(* Logix 5000 project; controller MV vendor 1 type 14 code 217 rev 31.11; software revision 31.00; part 48 of 53 *)
(* tags used below, declared in another part *)
   CWD : CHECKWORD_FLAGS;
   Delphi_Does_Eng_Func : BOOL;
   MV_MV1R : PlantItem;   // MV1R
   MV_MV20_CV1 : PlantItem;   // MV20_CV1
   MV_MV21_CV1 : PlantItem;   // MV21_CV1
   MV_MV22_CV1 : PlantItem;   // MV22_CV1
   MV_MV23_CV1 : PlantItem;   // MV23_CV1
   MV_MV2R : PlantItem;   // MV2R
   MV_MV35_CV1 : PlantItem;   // MV35_CV1
   MV_MV36_AV01 : PlantItem;   // MV36_AV01
   MV_MV37_AV01 : PlantItem;   // MV37_AV01
   MV_MV38_AV01 : PlantItem;   // MV38_AV01
   MV_MV39_AV01 : PlantItem;   // MV39_AV01
   MV_MV3R : PlantItem;   // MV3R
   MV_MV40_AV01 : PlantItem;   // MV40_AV01
   MV_MV41_AV01 : PlantItem;   // MV41_AV01
   MV_MV42_AV01 : PlantItem;   // MV42_AV01
   MV_MV43_AV01 : PlantItem;   // MV43_AV01
   MV_MV44_AV01 : PlantItem;   // MV44_AV01
   MV_MV45_AV01 : PlantItem;   // MV45_AV01
   MV_MV46_AV01 : PlantItem;   // MV46_AV01
   MV_MV47_AV01 : PlantItem;   // MV47_AV01
   MV_MV4R : PlantItem;   // MV4R
   MV_MV5R : PlantItem;   // MV5R
   MV_MV6R : PlantItem;   // MV6R
   MV_MV7R : PlantItem;   // MV7R
   MV_N255 : DINT[255];   // Old Format Checkwords To Keep Delphi Indicating Status Correctly.
(* MV_Common, continued *)

   24: [XIC(Delphi_Does_Eng_Func) [[XIC(MV_N255[24].8) [OTL(MV_MV35_CV1.CW.[CWD.MANUAL]) ,XIC(MV_N255[24].9) OTL(MV_MV35_CV1.CW.[CWD.MANDRV]) ,XIO(MV_N255[24].9) OTU(MV_MV35_CV1.CW.[CWD.MANDRV]) ] ,XIO(MV_N255[24].8) [OTU(MV_MV35_CV1.CW.[CWD.MANUAL]) ,[XIC(MV_MV35_CV1.CW.[CWD.OUTPUT]) OTL(MV_N255[24].9) ,XIO(MV_MV35_CV1.CW.[CWD.OUTPUT]) OTU(MV_N255[24].9) ] ] ] ,[XIC(MV_N255[24].13) OTL(MV_MV35_CV1.CW.[CWD.CHECKOFF]) ,XIO(MV_N255[24].13) OTU(MV_MV35_CV1.CW.[CWD.CHECKOFF]) ] ] ,XIO(Delphi_Does_Eng_Func) [[XIC(MV_MV35_CV1.CW.[CWD.MANUAL]) OTL(MV_N255[24].8) ,XIO(MV_MV35_CV1.CW.[CWD.MANUAL]) OTU(MV_N255[24].8) ] ,[XIC(MV_MV35_CV1.CW.[CWD.CHECKOFF]) OTL(MV_N255[24].13) ,XIO(MV_MV35_CV1.CW.[CWD.CHECKOFF]) OTU(MV_N255[24].13) ] ,[XIC(MV_MV35_CV1.CW.[CWD.OUTPUT]) OTL(MV_N255[24].9) ,XIO(MV_MV35_CV1.CW.[CWD.OUTPUT]) OTU(MV_N255[24].9) ] ] ,XIC(MV_MV35_CV1.CW.[CWD.OUTPUT]) OTE(MV_N255[24].10) ,XIO(MV_MV35_CV1.CW.[CWD.OUTPUT]) OTE(MV_N255[24].11) ,XIC(MV_MV35_CV1.CW.[CWD.FAULT]) OTE(MV_N255[24].15) ];
   25: [XIC(Delphi_Does_Eng_Func) [[XIC(MV_N255[25].8) [OTL(MV_MV20_CV1.CW.[CWD.MANUAL]) ,XIC(MV_N255[25].9) OTL(MV_MV20_CV1.CW.[CWD.MANDRV]) ,XIO(MV_N255[25].9) OTU(MV_MV20_CV1.CW.[CWD.MANDRV]) ] ,XIO(MV_N255[25].8) [OTU(MV_MV20_CV1.CW.[CWD.MANUAL]) ,[XIC(MV_MV20_CV1.CW.[CWD.OUTPUT]) OTL(MV_N255[25].9) ,XIO(MV_MV20_CV1.CW.[CWD.OUTPUT]) OTU(MV_N255[25].9) ] ] ] ,[XIC(MV_N255[25].13) OTL(MV_MV20_CV1.CW.[CWD.CHECKOFF]) ,XIO(MV_N255[25].13) OTU(MV_MV20_CV1.CW.[CWD.CHECKOFF]) ] ] ,XIO(Delphi_Does_Eng_Func) [[XIC(MV_MV20_CV1.CW.[CWD.MANUAL]) OTL(MV_N255[25].8) ,XIO(MV_MV20_CV1.CW.[CWD.MANUAL]) OTU(MV_N255[25].8) ] ,[XIC(MV_MV20_CV1.CW.[CWD.CHECKOFF]) OTL(MV_N255[25].13) ,XIO(MV_MV20_CV1.CW.[CWD.CHECKOFF]) OTU(MV_N255[25].13) ] ,[XIC(MV_MV20_CV1.CW.[CWD.OUTPUT]) OTL(MV_N255[25].9) ,XIO(MV_MV20_CV1.CW.[CWD.OUTPUT]) OTU(MV_N255[25].9) ] ] ,XIC(MV_MV20_CV1.CW.[CWD.OUTPUT]) OTE(MV_N255[25].10) ,XIO(MV_MV20_CV1.CW.[CWD.OUTPUT]) OTE(MV_N255[25].11) ,XIC(MV_MV20_CV1.CW.[CWD.FAULT]) OTE(MV_N255[25].15) ];
   26: [XIC(Delphi_Does_Eng_Func) [[XIC(MV_N255[26].8) [OTL(MV_MV21_CV1.CW.[CWD.MANUAL]) ,XIC(MV_N255[26].9) OTL(MV_MV21_CV1.CW.[CWD.MANDRV]) ,XIO(MV_N255[26].9) OTU(MV_MV21_CV1.CW.[CWD.MANDRV]) ] ,XIO(MV_N255[26].8) [OTU(MV_MV21_CV1.CW.[CWD.MANUAL]) ,[XIC(MV_MV21_CV1.CW.[CWD.OUTPUT]) OTL(MV_N255[26].9) ,XIO(MV_MV21_CV1.CW.[CWD.OUTPUT]) OTU(MV_N255[26].9) ] ] ] ,[XIC(MV_N255[26].13) OTL(MV_MV21_CV1.CW.[CWD.CHECKOFF]) ,XIO(MV_N255[26].13) OTU(MV_MV21_CV1.CW.[CWD.CHECKOFF]) ] ] ,XIO(Delphi_Does_Eng_Func) [[XIC(MV_MV21_CV1.CW.[CWD.MANUAL]) OTL(MV_N255[26].8) ,XIO(MV_MV21_CV1.CW.[CWD.MANUAL]) OTU(MV_N255[26].8) ] ,[XIC(MV_MV21_CV1.CW.[CWD.CHECKOFF]) OTL(MV_N255[26].13) ,XIO(MV_MV21_CV1.CW.[CWD.CHECKOFF]) OTU(MV_N255[26].13) ] ,[XIC(MV_MV21_CV1.CW.[CWD.OUTPUT]) OTL(MV_N255[26].9) ,XIO(MV_MV21_CV1.CW.[CWD.OUTPUT]) OTU(MV_N255[26].9) ] ] ,XIC(MV_MV21_CV1.CW.[CWD.OUTPUT]) OTE(MV_N255[26].10) ,XIO(MV_MV21_CV1.CW.[CWD.OUTPUT]) OTE(MV_N255[26].11) ,XIC(MV_MV21_CV1.CW.[CWD.FAULT]) OTE(MV_N255[26].15) ];
   27: [XIC(Delphi_Does_Eng_Func) [[XIC(MV_N255[27].8) [OTL(MV_MV22_CV1.CW.[CWD.MANUAL]) ,XIC(MV_N255[27].9) OTL(MV_MV22_CV1.CW.[CWD.MANDRV]) ,XIO(MV_N255[27].9) OTU(MV_MV22_CV1.CW.[CWD.MANDRV]) ] ,XIO(MV_N255[27].8) [OTU(MV_MV22_CV1.CW.[CWD.MANUAL]) ,[XIC(MV_MV22_CV1.CW.[CWD.OUTPUT]) OTL(MV_N255[27].9) ,XIO(MV_MV22_CV1.CW.[CWD.OUTPUT]) OTU(MV_N255[27].9) ] ] ] ,[XIC(MV_N255[27].13) OTL(MV_MV22_CV1.CW.[CWD.CHECKOFF]) ,XIO(MV_N255[27].13) OTU(MV_MV22_CV1.CW.[CWD.CHECKOFF]) ] ] ,XIO(Delphi_Does_Eng_Func) [[XIC(MV_MV22_CV1.CW.[CWD.MANUAL]) OTL(MV_N255[27].8) ,XIO(MV_MV22_CV1.CW.[CWD.MANUAL]) OTU(MV_N255[27].8) ] ,[XIC(MV_MV22_CV1.CW.[CWD.CHECKOFF]) OTL(MV_N255[27].13) ,XIO(MV_MV22_CV1.CW.[CWD.CHECKOFF]) OTU(MV_N255[27].13) ] ,[XIC(MV_MV22_CV1.CW.[CWD.OUTPUT]) OTL(MV_N255[27].9) ,XIO(MV_MV22_CV1.CW.[CWD.OUTPUT]) OTU(MV_N255[27].9) ] ] ,XIC(MV_MV22_CV1.CW.[CWD.OUTPUT]) OTE(MV_N255[27].10) ,XIO(MV_MV22_CV1.CW.[CWD.OUTPUT]) OTE(MV_N255[27].11) ,XIC(MV_MV22_CV1.CW.[CWD.FAULT]) OTE(MV_N255[27].15) ];
   28: [XIC(Delphi_Does_Eng_Func) [[XIC(MV_N255[28].8) [OTL(MV_MV23_CV1.CW.[CWD.MANUAL]) ,XIC(MV_N255[28].9) OTL(MV_MV23_CV1.CW.[CWD.MANDRV]) ,XIO(MV_N255[28].9) OTU(MV_MV23_CV1.CW.[CWD.MANDRV]) ] ,XIO(MV_N255[28].8) [OTU(MV_MV23_CV1.CW.[CWD.MANUAL]) ,[XIC(MV_MV23_CV1.CW.[CWD.OUTPUT]) OTL(MV_N255[28].9) ,XIO(MV_MV23_CV1.CW.[CWD.OUTPUT]) OTU(MV_N255[28].9) ] ] ] ,[XIC(MV_N255[28].13) OTL(MV_MV23_CV1.CW.[CWD.CHECKOFF]) ,XIO(MV_N255[28].13) OTU(MV_MV23_CV1.CW.[CWD.CHECKOFF]) ] ] ,XIO(Delphi_Does_Eng_Func) [[XIC(MV_MV23_CV1.CW.[CWD.MANUAL]) OTL(MV_N255[28].8) ,XIO(MV_MV23_CV1.CW.[CWD.MANUAL]) OTU(MV_N255[28].8) ] ,[XIC(MV_MV23_CV1.CW.[CWD.CHECKOFF]) OTL(MV_N255[28].13) ,XIO(MV_MV23_CV1.CW.[CWD.CHECKOFF]) OTU(MV_N255[28].13) ] ,[XIC(MV_MV23_CV1.CW.[CWD.OUTPUT]) OTL(MV_N255[28].9) ,XIO(MV_MV23_CV1.CW.[CWD.OUTPUT]) OTU(MV_N255[28].9) ] ] ,XIC(MV_MV23_CV1.CW.[CWD.OUTPUT]) OTE(MV_N255[28].10) ,XIO(MV_MV23_CV1.CW.[CWD.OUTPUT]) OTE(MV_N255[28].11) ,XIC(MV_MV23_CV1.CW.[CWD.FAULT]) OTE(MV_N255[28].15) ];
   29: [XIC(Delphi_Does_Eng_Func) [[XIC(MV_N255[64].8) [OTL(MV_MV36_AV01.CW.[CWD.MANUAL]) ,XIC(MV_N255[64].9) OTL(MV_MV36_AV01.CW.[CWD.MANDRV]) ,XIO(MV_N255[64].9) OTU(MV_MV36_AV01.CW.[CWD.MANDRV]) ] ,XIO(MV_N255[64].8) [OTU(MV_MV36_AV01.CW.[CWD.MANUAL]) ,[XIC(MV_MV36_AV01.CW.[CWD.OUTPUT]) OTL(MV_N255[64].9) ,XIO(MV_MV36_AV01.CW.[CWD.OUTPUT]) OTU(MV_N255[64].9) ] ] ] ,[XIC(MV_N255[64].13) OTL(MV_MV36_AV01.CW.[CWD.CHECKOFF]) ,XIO(MV_N255[64].13) OTU(MV_MV36_AV01.CW.[CWD.CHECKOFF]) ] ] ,XIO(Delphi_Does_Eng_Func) [[XIC(MV_MV36_AV01.CW.[CWD.MANUAL]) OTL(MV_N255[64].8) ,XIO(MV_MV36_AV01.CW.[CWD.MANUAL]) OTU(MV_N255[64].8) ] ,[XIC(MV_MV36_AV01.CW.[CWD.CHECKOFF]) OTL(MV_N255[64].13) ,XIO(MV_MV36_AV01.CW.[CWD.CHECKOFF]) OTU(MV_N255[64].13) ] ,[XIC(MV_MV36_AV01.CW.[CWD.OUTPUT]) OTL(MV_N255[64].9) ,XIO(MV_MV36_AV01.CW.[CWD.OUTPUT]) OTU(MV_N255[64].9) ] ] ,XIC(MV_MV36_AV01.CW.[CWD.OUTPUT]) OTE(MV_N255[64].10) ,XIO(MV_MV36_AV01.CW.[CWD.OUTPUT]) OTE(MV_N255[64].11) ,XIC(MV_MV36_AV01.CW.[CWD.FAULT]) OTE(MV_N255[64].15) ];
   30: [XIC(Delphi_Does_Eng_Func) [[XIC(MV_N255[65].8) [OTL(MV_MV37_AV01.CW.[CWD.MANUAL]) ,XIC(MV_N255[65].9) OTL(MV_MV37_AV01.CW.[CWD.MANDRV]) ,XIO(MV_N255[65].9) OTU(MV_MV37_AV01.CW.[CWD.MANDRV]) ] ,XIO(MV_N255[65].8) [OTU(MV_MV37_AV01.CW.[CWD.MANUAL]) ,[XIC(MV_MV37_AV01.CW.[CWD.OUTPUT]) OTL(MV_N255[65].9) ,XIO(MV_MV37_AV01.CW.[CWD.OUTPUT]) OTU(MV_N255[65].9) ] ] ] ,[XIC(MV_N255[65].13) OTL(MV_MV37_AV01.CW.[CWD.CHECKOFF]) ,XIO(MV_N255[65].13) OTU(MV_MV37_AV01.CW.[CWD.CHECKOFF]) ] ] ,XIO(Delphi_Does_Eng_Func) [[XIC(MV_MV37_AV01.CW.[CWD.MANUAL]) OTL(MV_N255[65].8) ,XIO(MV_MV37_AV01.CW.[CWD.MANUAL]) OTU(MV_N255[65].8) ] ,[XIC(MV_MV37_AV01.CW.[CWD.CHECKOFF]) OTL(MV_N255[65].13) ,XIO(MV_MV37_AV01.CW.[CWD.CHECKOFF]) OTU(MV_N255[65].13) ] ,[XIC(MV_MV37_AV01.CW.[CWD.OUTPUT]) OTL(MV_N255[65].9) ,XIO(MV_MV37_AV01.CW.[CWD.OUTPUT]) OTU(MV_N255[65].9) ] ] ,XIC(MV_MV37_AV01.CW.[CWD.OUTPUT]) OTE(MV_N255[65].10) ,XIO(MV_MV37_AV01.CW.[CWD.OUTPUT]) OTE(MV_N255[65].11) ,XIC(MV_MV37_AV01.CW.[CWD.FAULT]) OTE(MV_N255[65].15) ];
   31: [XIC(Delphi_Does_Eng_Func) [[XIC(MV_N255[66].8) [OTL(MV_MV38_AV01.CW.[CWD.MANUAL]) ,XIC(MV_N255[66].9) OTL(MV_MV38_AV01.CW.[CWD.MANDRV]) ,XIO(MV_N255[66].9) OTU(MV_MV38_AV01.CW.[CWD.MANDRV]) ] ,XIO(MV_N255[66].8) [OTU(MV_MV38_AV01.CW.[CWD.MANUAL]) ,[XIC(MV_MV38_AV01.CW.[CWD.OUTPUT]) OTL(MV_N255[66].9) ,XIO(MV_MV38_AV01.CW.[CWD.OUTPUT]) OTU(MV_N255[66].9) ] ] ] ,[XIC(MV_N255[66].13) OTL(MV_MV38_AV01.CW.[CWD.CHECKOFF]) ,XIO(MV_N255[66].13) OTU(MV_MV38_AV01.CW.[CWD.CHECKOFF]) ] ] ,XIO(Delphi_Does_Eng_Func) [[XIC(MV_MV38_AV01.CW.[CWD.MANUAL]) OTL(MV_N255[66].8) ,XIO(MV_MV38_AV01.CW.[CWD.MANUAL]) OTU(MV_N255[66].8) ] ,[XIC(MV_MV38_AV01.CW.[CWD.CHECKOFF]) OTL(MV_N255[66].13) ,XIO(MV_MV38_AV01.CW.[CWD.CHECKOFF]) OTU(MV_N255[66].13) ] ,[XIC(MV_MV38_AV01.CW.[CWD.OUTPUT]) OTL(MV_N255[66].9) ,XIO(MV_MV38_AV01.CW.[CWD.OUTPUT]) OTU(MV_N255[66].9) ] ] ,XIC(MV_MV38_AV01.CW.[CWD.OUTPUT]) OTE(MV_N255[66].10) ,XIO(MV_MV38_AV01.CW.[CWD.OUTPUT]) OTE(MV_N255[66].11) ,XIC(MV_MV38_AV01.CW.[CWD.FAULT]) OTE(MV_N255[66].15) ];
   32: [XIC(Delphi_Does_Eng_Func) [[XIC(MV_N255[67].8) [OTL(MV_MV39_AV01.CW.[CWD.MANUAL]) ,XIC(MV_N255[67].9) OTL(MV_MV39_AV01.CW.[CWD.MANDRV]) ,XIO(MV_N255[67].9) OTU(MV_MV39_AV01.CW.[CWD.MANDRV]) ] ,XIO(MV_N255[67].8) [OTU(MV_MV39_AV01.CW.[CWD.MANUAL]) ,[XIC(MV_MV39_AV01.CW.[CWD.OUTPUT]) OTL(MV_N255[67].9) ,XIO(MV_MV39_AV01.CW.[CWD.OUTPUT]) OTU(MV_N255[67].9) ] ] ] ,[XIC(MV_N255[67].13) OTL(MV_MV39_AV01.CW.[CWD.CHECKOFF]) ,XIO(MV_N255[67].13) OTU(MV_MV39_AV01.CW.[CWD.CHECKOFF]) ] ] ,XIO(Delphi_Does_Eng_Func) [[XIC(MV_MV39_AV01.CW.[CWD.MANUAL]) OTL(MV_N255[67].8) ,XIO(MV_MV39_AV01.CW.[CWD.MANUAL]) OTU(MV_N255[67].8) ] ,[XIC(MV_MV39_AV01.CW.[CWD.CHECKOFF]) OTL(MV_N255[67].13) ,XIO(MV_MV39_AV01.CW.[CWD.CHECKOFF]) OTU(MV_N255[67].13) ] ,[XIC(MV_MV39_AV01.CW.[CWD.OUTPUT]) OTL(MV_N255[67].9) ,XIO(MV_MV39_AV01.CW.[CWD.OUTPUT]) OTU(MV_N255[67].9) ] ] ,XIC(MV_MV39_AV01.CW.[CWD.OUTPUT]) OTE(MV_N255[67].10) ,XIO(MV_MV39_AV01.CW.[CWD.OUTPUT]) OTE(MV_N255[67].11) ,XIC(MV_MV39_AV01.CW.[CWD.FAULT]) OTE(MV_N255[67].15) ];
   33: [XIC(Delphi_Does_Eng_Func) [[XIC(MV_N255[68].8) [OTL(MV_MV40_AV01.CW.[CWD.MANUAL]) ,XIC(MV_N255[68].9) OTL(MV_MV40_AV01.CW.[CWD.MANDRV]) ,XIO(MV_N255[68].9) OTU(MV_MV40_AV01.CW.[CWD.MANDRV]) ] ,XIO(MV_N255[68].8) [OTU(MV_MV40_AV01.CW.[CWD.MANUAL]) ,[XIC(MV_MV40_AV01.CW.[CWD.OUTPUT]) OTL(MV_N255[68].9) ,XIO(MV_MV40_AV01.CW.[CWD.OUTPUT]) OTU(MV_N255[68].9) ] ] ] ,[XIC(MV_N255[68].13) OTL(MV_MV40_AV01.CW.[CWD.CHECKOFF]) ,XIO(MV_N255[68].13) OTU(MV_MV40_AV01.CW.[CWD.CHECKOFF]) ] ] ,XIO(Delphi_Does_Eng_Func) [[XIC(MV_MV40_AV01.CW.[CWD.MANUAL]) OTL(MV_N255[68].8) ,XIO(MV_MV40_AV01.CW.[CWD.MANUAL]) OTU(MV_N255[68].8) ] ,[XIC(MV_MV40_AV01.CW.[CWD.CHECKOFF]) OTL(MV_N255[68].13) ,XIO(MV_MV40_AV01.CW.[CWD.CHECKOFF]) OTU(MV_N255[68].13) ] ,[XIC(MV_MV40_AV01.CW.[CWD.OUTPUT]) OTL(MV_N255[68].9) ,XIO(MV_MV40_AV01.CW.[CWD.OUTPUT]) OTU(MV_N255[68].9) ] ] ,XIC(MV_MV40_AV01.CW.[CWD.OUTPUT]) OTE(MV_N255[68].10) ,XIO(MV_MV40_AV01.CW.[CWD.OUTPUT]) OTE(MV_N255[68].11) ,XIC(MV_MV40_AV01.CW.[CWD.FAULT]) OTE(MV_N255[68].15) ];
   34: [XIC(Delphi_Does_Eng_Func) [[XIC(MV_N255[69].8) [OTL(MV_MV41_AV01.CW.[CWD.MANUAL]) ,XIC(MV_N255[69].9) OTL(MV_MV41_AV01.CW.[CWD.MANDRV]) ,XIO(MV_N255[69].9) OTU(MV_MV41_AV01.CW.[CWD.MANDRV]) ] ,XIO(MV_N255[69].8) [OTU(MV_MV41_AV01.CW.[CWD.MANUAL]) ,[XIC(MV_MV41_AV01.CW.[CWD.OUTPUT]) OTL(MV_N255[69].9) ,XIO(MV_MV41_AV01.CW.[CWD.OUTPUT]) OTU(MV_N255[69].9) ] ] ] ,[XIC(MV_N255[69].13) OTL(MV_MV41_AV01.CW.[CWD.CHECKOFF]) ,XIO(MV_N255[69].13) OTU(MV_MV41_AV01.CW.[CWD.CHECKOFF]) ] ] ,XIO(Delphi_Does_Eng_Func) [[XIC(MV_MV41_AV01.CW.[CWD.MANUAL]) OTL(MV_N255[69].8) ,XIO(MV_MV41_AV01.CW.[CWD.MANUAL]) OTU(MV_N255[69].8) ] ,[XIC(MV_MV41_AV01.CW.[CWD.CHECKOFF]) OTL(MV_N255[69].13) ,XIO(MV_MV41_AV01.CW.[CWD.CHECKOFF]) OTU(MV_N255[69].13) ] ,[XIC(MV_MV41_AV01.CW.[CWD.OUTPUT]) OTL(MV_N255[69].9) ,XIO(MV_MV41_AV01.CW.[CWD.OUTPUT]) OTU(MV_N255[69].9) ] ] ,XIC(MV_MV41_AV01.CW.[CWD.OUTPUT]) OTE(MV_N255[69].10) ,XIO(MV_MV41_AV01.CW.[CWD.OUTPUT]) OTE(MV_N255[69].11) ,XIC(MV_MV41_AV01.CW.[CWD.FAULT]) OTE(MV_N255[69].15) ];
   35: [XIC(Delphi_Does_Eng_Func) [[XIC(MV_N255[70].8) [OTL(MV_MV42_AV01.CW.[CWD.MANUAL]) ,XIC(MV_N255[70].9) OTL(MV_MV42_AV01.CW.[CWD.MANDRV]) ,XIO(MV_N255[70].9) OTU(MV_MV42_AV01.CW.[CWD.MANDRV]) ] ,XIO(MV_N255[70].8) [OTU(MV_MV42_AV01.CW.[CWD.MANUAL]) ,[XIC(MV_MV42_AV01.CW.[CWD.OUTPUT]) OTL(MV_N255[70].9) ,XIO(MV_MV42_AV01.CW.[CWD.OUTPUT]) OTU(MV_N255[70].9) ] ] ] ,[XIC(MV_N255[70].13) OTL(MV_MV42_AV01.CW.[CWD.CHECKOFF]) ,XIO(MV_N255[70].13) OTU(MV_MV42_AV01.CW.[CWD.CHECKOFF]) ] ] ,XIO(Delphi_Does_Eng_Func) [[XIC(MV_MV42_AV01.CW.[CWD.MANUAL]) OTL(MV_N255[70].8) ,XIO(MV_MV42_AV01.CW.[CWD.MANUAL]) OTU(MV_N255[70].8) ] ,[XIC(MV_MV42_AV01.CW.[CWD.CHECKOFF]) OTL(MV_N255[70].13) ,XIO(MV_MV42_AV01.CW.[CWD.CHECKOFF]) OTU(MV_N255[70].13) ] ,[XIC(MV_MV42_AV01.CW.[CWD.OUTPUT]) OTL(MV_N255[70].9) ,XIO(MV_MV42_AV01.CW.[CWD.OUTPUT]) OTU(MV_N255[70].9) ] ] ,XIC(MV_MV42_AV01.CW.[CWD.OUTPUT]) OTE(MV_N255[70].10) ,XIO(MV_MV42_AV01.CW.[CWD.OUTPUT]) OTE(MV_N255[70].11) ,XIC(MV_MV42_AV01.CW.[CWD.FAULT]) OTE(MV_N255[70].15) ];
   36: [XIC(Delphi_Does_Eng_Func) [[XIC(MV_N255[71].8) [OTL(MV_MV43_AV01.CW.[CWD.MANUAL]) ,XIC(MV_N255[71].9) OTL(MV_MV43_AV01.CW.[CWD.MANDRV]) ,XIO(MV_N255[71].9) OTU(MV_MV43_AV01.CW.[CWD.MANDRV]) ] ,XIO(MV_N255[71].8) [OTU(MV_MV43_AV01.CW.[CWD.MANUAL]) ,[XIC(MV_MV43_AV01.CW.[CWD.OUTPUT]) OTL(MV_N255[71].9) ,XIO(MV_MV43_AV01.CW.[CWD.OUTPUT]) OTU(MV_N255[71].9) ] ] ] ,[XIC(MV_N255[71].13) OTL(MV_MV43_AV01.CW.[CWD.CHECKOFF]) ,XIO(MV_N255[71].13) OTU(MV_MV43_AV01.CW.[CWD.CHECKOFF]) ] ] ,XIO(Delphi_Does_Eng_Func) [[XIC(MV_MV43_AV01.CW.[CWD.MANUAL]) OTL(MV_N255[71].8) ,XIO(MV_MV43_AV01.CW.[CWD.MANUAL]) OTU(MV_N255[71].8) ] ,[XIC(MV_MV43_AV01.CW.[CWD.CHECKOFF]) OTL(MV_N255[71].13) ,XIO(MV_MV43_AV01.CW.[CWD.CHECKOFF]) OTU(MV_N255[71].13) ] ,[XIC(MV_MV43_AV01.CW.[CWD.OUTPUT]) OTL(MV_N255[71].9) ,XIO(MV_MV43_AV01.CW.[CWD.OUTPUT]) OTU(MV_N255[71].9) ] ] ,XIC(MV_MV43_AV01.CW.[CWD.OUTPUT]) OTE(MV_N255[71].10) ,XIO(MV_MV43_AV01.CW.[CWD.OUTPUT]) OTE(MV_N255[71].11) ,XIC(MV_MV43_AV01.CW.[CWD.FAULT]) OTE(MV_N255[71].15) ];
   37: [XIC(Delphi_Does_Eng_Func) [[XIC(MV_N255[72].8) [OTL(MV_MV44_AV01.CW.[CWD.MANUAL]) ,XIC(MV_N255[72].9) OTL(MV_MV44_AV01.CW.[CWD.MANDRV]) ,XIO(MV_N255[72].9) OTU(MV_MV44_AV01.CW.[CWD.MANDRV]) ] ,XIO(MV_N255[72].8) [OTU(MV_MV44_AV01.CW.[CWD.MANUAL]) ,[XIC(MV_MV44_AV01.CW.[CWD.OUTPUT]) OTL(MV_N255[72].9) ,XIO(MV_MV44_AV01.CW.[CWD.OUTPUT]) OTU(MV_N255[72].9) ] ] ] ,[XIC(MV_N255[72].13) OTL(MV_MV44_AV01.CW.[CWD.CHECKOFF]) ,XIO(MV_N255[72].13) OTU(MV_MV44_AV01.CW.[CWD.CHECKOFF]) ] ] ,XIO(Delphi_Does_Eng_Func) [[XIC(MV_MV44_AV01.CW.[CWD.MANUAL]) OTL(MV_N255[72].8) ,XIO(MV_MV44_AV01.CW.[CWD.MANUAL]) OTU(MV_N255[72].8) ] ,[XIC(MV_MV44_AV01.CW.[CWD.CHECKOFF]) OTL(MV_N255[72].13) ,XIO(MV_MV44_AV01.CW.[CWD.CHECKOFF]) OTU(MV_N255[72].13) ] ,[XIC(MV_MV44_AV01.CW.[CWD.OUTPUT]) OTL(MV_N255[72].9) ,XIO(MV_MV44_AV01.CW.[CWD.OUTPUT]) OTU(MV_N255[72].9) ] ] ,XIC(MV_MV44_AV01.CW.[CWD.OUTPUT]) OTE(MV_N255[72].10) ,XIO(MV_MV44_AV01.CW.[CWD.OUTPUT]) OTE(MV_N255[72].11) ,XIC(MV_MV44_AV01.CW.[CWD.FAULT]) OTE(MV_N255[72].15) ];
   38: [XIC(Delphi_Does_Eng_Func) [[XIC(MV_N255[73].8) [OTL(MV_MV45_AV01.CW.[CWD.MANUAL]) ,XIC(MV_N255[73].9) OTL(MV_MV45_AV01.CW.[CWD.MANDRV]) ,XIO(MV_N255[73].9) OTU(MV_MV45_AV01.CW.[CWD.MANDRV]) ] ,XIO(MV_N255[73].8) [OTU(MV_MV45_AV01.CW.[CWD.MANUAL]) ,[XIC(MV_MV45_AV01.CW.[CWD.OUTPUT]) OTL(MV_N255[73].9) ,XIO(MV_MV45_AV01.CW.[CWD.OUTPUT]) OTU(MV_N255[73].9) ] ] ] ,[XIC(MV_N255[73].13) OTL(MV_MV45_AV01.CW.[CWD.CHECKOFF]) ,XIO(MV_N255[73].13) OTU(MV_MV45_AV01.CW.[CWD.CHECKOFF]) ] ] ,XIO(Delphi_Does_Eng_Func) [[XIC(MV_MV45_AV01.CW.[CWD.MANUAL]) OTL(MV_N255[73].8) ,XIO(MV_MV45_AV01.CW.[CWD.MANUAL]) OTU(MV_N255[73].8) ] ,[XIC(MV_MV45_AV01.CW.[CWD.CHECKOFF]) OTL(MV_N255[73].13) ,XIO(MV_MV45_AV01.CW.[CWD.CHECKOFF]) OTU(MV_N255[73].13) ] ,[XIC(MV_MV45_AV01.CW.[CWD.OUTPUT]) OTL(MV_N255[73].9) ,XIO(MV_MV45_AV01.CW.[CWD.OUTPUT]) OTU(MV_N255[73].9) ] ] ,XIC(MV_MV45_AV01.CW.[CWD.OUTPUT]) OTE(MV_N255[73].10) ,XIO(MV_MV45_AV01.CW.[CWD.OUTPUT]) OTE(MV_N255[73].11) ,XIC(MV_MV45_AV01.CW.[CWD.FAULT]) OTE(MV_N255[73].15) ];
   39: [XIC(Delphi_Does_Eng_Func) [[XIC(MV_N255[74].8) [OTL(MV_MV46_AV01.CW.[CWD.MANUAL]) ,XIC(MV_N255[74].9) OTL(MV_MV46_AV01.CW.[CWD.MANDRV]) ,XIO(MV_N255[74].9) OTU(MV_MV46_AV01.CW.[CWD.MANDRV]) ] ,XIO(MV_N255[74].8) [OTU(MV_MV46_AV01.CW.[CWD.MANUAL]) ,[XIC(MV_MV46_AV01.CW.[CWD.OUTPUT]) OTL(MV_N255[74].9) ,XIO(MV_MV46_AV01.CW.[CWD.OUTPUT]) OTU(MV_N255[74].9) ] ] ] ,[XIC(MV_N255[74].13) OTL(MV_MV46_AV01.CW.[CWD.CHECKOFF]) ,XIO(MV_N255[74].13) OTU(MV_MV46_AV01.CW.[CWD.CHECKOFF]) ] ] ,XIO(Delphi_Does_Eng_Func) [[XIC(MV_MV46_AV01.CW.[CWD.MANUAL]) OTL(MV_N255[74].8) ,XIO(MV_MV46_AV01.CW.[CWD.MANUAL]) OTU(MV_N255[74].8) ] ,[XIC(MV_MV46_AV01.CW.[CWD.CHECKOFF]) OTL(MV_N255[74].13) ,XIO(MV_MV46_AV01.CW.[CWD.CHECKOFF]) OTU(MV_N255[74].13) ] ,[XIC(MV_MV46_AV01.CW.[CWD.OUTPUT]) OTL(MV_N255[74].9) ,XIO(MV_MV46_AV01.CW.[CWD.OUTPUT]) OTU(MV_N255[74].9) ] ] ,XIC(MV_MV46_AV01.CW.[CWD.OUTPUT]) OTE(MV_N255[74].10) ,XIO(MV_MV46_AV01.CW.[CWD.OUTPUT]) OTE(MV_N255[74].11) ,XIC(MV_MV46_AV01.CW.[CWD.FAULT]) OTE(MV_N255[74].15) ];
   40: [XIC(Delphi_Does_Eng_Func) [[XIC(MV_N255[75].8) [OTL(MV_MV47_AV01.CW.[CWD.MANUAL]) ,XIC(MV_N255[75].9) OTL(MV_MV47_AV01.CW.[CWD.MANDRV]) ,XIO(MV_N255[75].9) OTU(MV_MV47_AV01.CW.[CWD.MANDRV]) ] ,XIO(MV_N255[75].8) [OTU(MV_MV47_AV01.CW.[CWD.MANUAL]) ,[XIC(MV_MV47_AV01.CW.[CWD.OUTPUT]) OTL(MV_N255[75].9) ,XIO(MV_MV47_AV01.CW.[CWD.OUTPUT]) OTU(MV_N255[75].9) ] ] ] ,[XIC(MV_N255[75].13) OTL(MV_MV47_AV01.CW.[CWD.CHECKOFF]) ,XIO(MV_N255[75].13) OTU(MV_MV47_AV01.CW.[CWD.CHECKOFF]) ] ] ,XIO(Delphi_Does_Eng_Func) [[XIC(MV_MV47_AV01.CW.[CWD.MANUAL]) OTL(MV_N255[75].8) ,XIO(MV_MV47_AV01.CW.[CWD.MANUAL]) OTU(MV_N255[75].8) ] ,[XIC(MV_MV47_AV01.CW.[CWD.CHECKOFF]) OTL(MV_N255[75].13) ,XIO(MV_MV47_AV01.CW.[CWD.CHECKOFF]) OTU(MV_N255[75].13) ] ,[XIC(MV_MV47_AV01.CW.[CWD.OUTPUT]) OTL(MV_N255[75].9) ,XIO(MV_MV47_AV01.CW.[CWD.OUTPUT]) OTU(MV_N255[75].9) ] ] ,XIC(MV_MV47_AV01.CW.[CWD.OUTPUT]) OTE(MV_N255[75].10) ,XIO(MV_MV47_AV01.CW.[CWD.OUTPUT]) OTE(MV_N255[75].11) ,XIC(MV_MV47_AV01.CW.[CWD.FAULT]) OTE(MV_N255[75].15) ];
   41: [XIC(Delphi_Does_Eng_Func) [[XIC(MV_N255[32].8) [OTL(MV_MV1R.CW.[CWD.MANUAL]) ,XIC(MV_N255[32].9) OTL(MV_MV1R.CW.[CWD.MANDRV]) ,XIO(MV_N255[32].9) OTU(MV_MV1R.CW.[CWD.MANDRV]) ] ,XIO(MV_N255[32].8) [OTU(MV_MV1R.CW.[CWD.MANUAL]) ,[XIC(MV_MV1R.CW.[CWD.OUTPUT]) OTL(MV_N255[32].9) ,XIO(MV_MV1R.CW.[CWD.OUTPUT]) OTU(MV_N255[32].9) ] ] ] ,[XIC(MV_N255[32].13) OTL(MV_MV1R.CW.[CWD.CHECKOFF]) ,XIO(MV_N255[32].13) OTU(MV_MV1R.CW.[CWD.CHECKOFF]) ] ] ,XIO(Delphi_Does_Eng_Func) [[XIC(MV_MV1R.CW.[CWD.MANUAL]) OTL(MV_N255[32].8) ,XIO(MV_MV1R.CW.[CWD.MANUAL]) OTU(MV_N255[32].8) ] ,[XIC(MV_MV1R.CW.[CWD.CHECKOFF]) OTL(MV_N255[32].13) ,XIO(MV_MV1R.CW.[CWD.CHECKOFF]) OTU(MV_N255[32].13) ] ,[XIC(MV_MV1R.CW.[CWD.OUTPUT]) OTL(MV_N255[32].9) ,XIO(MV_MV1R.CW.[CWD.OUTPUT]) OTU(MV_N255[32].9) ] ] ,XIC(MV_MV1R.CW.[CWD.RUNFB]) OTE(MV_N255[32].10) ,XIO(MV_MV1R.CW.[CWD.RUNFB]) OTE(MV_N255[32].11) ,XIC(MV_MV1R.CW.[CWD.FAULT]) OTE(MV_N255[32].15) ];
   42: [XIC(Delphi_Does_Eng_Func) [[XIC(MV_N255[33].8) [OTL(MV_MV2R.CW.[CWD.MANUAL]) ,XIC(MV_N255[33].9) OTL(MV_MV2R.CW.[CWD.MANDRV]) ,XIO(MV_N255[33].9) OTU(MV_MV2R.CW.[CWD.MANDRV]) ] ,XIO(MV_N255[33].8) [OTU(MV_MV2R.CW.[CWD.MANUAL]) ,[XIC(MV_MV2R.CW.[CWD.OUTPUT]) OTL(MV_N255[33].9) ,XIO(MV_MV2R.CW.[CWD.OUTPUT]) OTU(MV_N255[33].9) ] ] ] ,[XIC(MV_N255[33].13) OTL(MV_MV2R.CW.[CWD.CHECKOFF]) ,XIO(MV_N255[33].13) OTU(MV_MV2R.CW.[CWD.CHECKOFF]) ] ] ,XIO(Delphi_Does_Eng_Func) [[XIC(MV_MV2R.CW.[CWD.MANUAL]) OTL(MV_N255[33].8) ,XIO(MV_MV2R.CW.[CWD.MANUAL]) OTU(MV_N255[33].8) ] ,[XIC(MV_MV2R.CW.[CWD.CHECKOFF]) OTL(MV_N255[33].13) ,XIO(MV_MV2R.CW.[CWD.CHECKOFF]) OTU(MV_N255[33].13) ] ,[XIC(MV_MV2R.CW.[CWD.OUTPUT]) OTL(MV_N255[33].9) ,XIO(MV_MV2R.CW.[CWD.OUTPUT]) OTU(MV_N255[33].9) ] ] ,XIC(MV_MV2R.CW.[CWD.RUNFB]) OTE(MV_N255[33].10) ,XIO(MV_MV2R.CW.[CWD.RUNFB]) OTE(MV_N255[33].11) ,XIC(MV_MV2R.CW.[CWD.FAULT]) OTE(MV_N255[33].15) ];
   43: [XIC(Delphi_Does_Eng_Func) [[XIC(MV_N255[34].8) [OTL(MV_MV3R.CW.[CWD.MANUAL]) ,XIC(MV_N255[34].9) OTL(MV_MV3R.CW.[CWD.MANDRV]) ,XIO(MV_N255[34].9) OTU(MV_MV3R.CW.[CWD.MANDRV]) ] ,XIO(MV_N255[34].8) [OTU(MV_MV3R.CW.[CWD.MANUAL]) ,[XIC(MV_MV3R.CW.[CWD.OUTPUT]) OTL(MV_N255[34].9) ,XIO(MV_MV3R.CW.[CWD.OUTPUT]) OTU(MV_N255[34].9) ] ] ] ,[XIC(MV_N255[34].13) OTL(MV_MV3R.CW.[CWD.CHECKOFF]) ,XIO(MV_N255[34].13) OTU(MV_MV3R.CW.[CWD.CHECKOFF]) ] ] ,XIO(Delphi_Does_Eng_Func) [[XIC(MV_MV3R.CW.[CWD.MANUAL]) OTL(MV_N255[34].8) ,XIO(MV_MV3R.CW.[CWD.MANUAL]) OTU(MV_N255[34].8) ] ,[XIC(MV_MV3R.CW.[CWD.CHECKOFF]) OTL(MV_N255[34].13) ,XIO(MV_MV3R.CW.[CWD.CHECKOFF]) OTU(MV_N255[34].13) ] ,[XIC(MV_MV3R.CW.[CWD.OUTPUT]) OTL(MV_N255[34].9) ,XIO(MV_MV3R.CW.[CWD.OUTPUT]) OTU(MV_N255[34].9) ] ] ,XIC(MV_MV3R.CW.[CWD.RUNFB]) OTE(MV_N255[34].10) ,XIO(MV_MV3R.CW.[CWD.RUNFB]) OTE(MV_N255[34].11) ,XIC(MV_MV3R.CW.[CWD.FAULT]) OTE(MV_N255[34].15) ];
   44: [XIC(Delphi_Does_Eng_Func) [[XIC(MV_N255[35].8) [OTL(MV_MV4R.CW.[CWD.MANUAL]) ,XIC(MV_N255[35].9) OTL(MV_MV4R.CW.[CWD.MANDRV]) ,XIO(MV_N255[35].9) OTU(MV_MV4R.CW.[CWD.MANDRV]) ] ,XIO(MV_N255[35].8) [OTU(MV_MV4R.CW.[CWD.MANUAL]) ,[XIC(MV_MV4R.CW.[CWD.OUTPUT]) OTL(MV_N255[35].9) ,XIO(MV_MV4R.CW.[CWD.OUTPUT]) OTU(MV_N255[35].9) ] ] ] ,[XIC(MV_N255[35].13) OTL(MV_MV4R.CW.[CWD.CHECKOFF]) ,XIO(MV_N255[35].13) OTU(MV_MV4R.CW.[CWD.CHECKOFF]) ] ] ,XIO(Delphi_Does_Eng_Func) [[XIC(MV_MV4R.CW.[CWD.MANUAL]) OTL(MV_N255[35].8) ,XIO(MV_MV4R.CW.[CWD.MANUAL]) OTU(MV_N255[35].8) ] ,[XIC(MV_MV4R.CW.[CWD.CHECKOFF]) OTL(MV_N255[35].13) ,XIO(MV_MV4R.CW.[CWD.CHECKOFF]) OTU(MV_N255[35].13) ] ,[XIC(MV_MV4R.CW.[CWD.OUTPUT]) OTL(MV_N255[35].9) ,XIO(MV_MV4R.CW.[CWD.OUTPUT]) OTU(MV_N255[35].9) ] ] ,XIC(MV_MV4R.CW.[CWD.RUNFB]) OTE(MV_N255[35].10) ,XIO(MV_MV4R.CW.[CWD.RUNFB]) OTE(MV_N255[35].11) ,XIC(MV_MV4R.CW.[CWD.FAULT]) OTE(MV_N255[35].15) ];
   45: [XIC(Delphi_Does_Eng_Func) [[XIC(MV_N255[36].8) [OTL(MV_MV5R.CW.[CWD.MANUAL]) ,XIC(MV_N255[36].9) OTL(MV_MV5R.CW.[CWD.MANDRV]) ,XIO(MV_N255[36].9) OTU(MV_MV5R.CW.[CWD.MANDRV]) ] ,XIO(MV_N255[36].8) [OTU(MV_MV5R.CW.[CWD.MANUAL]) ,[XIC(MV_MV5R.CW.[CWD.OUTPUT]) OTL(MV_N255[36].9) ,XIO(MV_MV5R.CW.[CWD.OUTPUT]) OTU(MV_N255[36].9) ] ] ] ,[XIC(MV_N255[36].13) OTL(MV_MV5R.CW.[CWD.CHECKOFF]) ,XIO(MV_N255[36].13) OTU(MV_MV5R.CW.[CWD.CHECKOFF]) ] ] ,XIO(Delphi_Does_Eng_Func) [[XIC(MV_MV5R.CW.[CWD.MANUAL]) OTL(MV_N255[36].8) ,XIO(MV_MV5R.CW.[CWD.MANUAL]) OTU(MV_N255[36].8) ] ,[XIC(MV_MV5R.CW.[CWD.CHECKOFF]) OTL(MV_N255[36].13) ,XIO(MV_MV5R.CW.[CWD.CHECKOFF]) OTU(MV_N255[36].13) ] ,[XIC(MV_MV5R.CW.[CWD.OUTPUT]) OTL(MV_N255[36].9) ,XIO(MV_MV5R.CW.[CWD.OUTPUT]) OTU(MV_N255[36].9) ] ] ,XIC(MV_MV5R.CW.[CWD.RUNFB]) OTE(MV_N255[36].10) ,XIO(MV_MV5R.CW.[CWD.RUNFB]) OTE(MV_N255[36].11) ,XIC(MV_MV5R.CW.[CWD.FAULT]) OTE(MV_N255[36].15) ];
   46: [XIC(Delphi_Does_Eng_Func) [[XIC(MV_N255[37].8) [OTL(MV_MV6R.CW.[CWD.MANUAL]) ,XIC(MV_N255[37].9) OTL(MV_MV6R.CW.[CWD.MANDRV]) ,XIO(MV_N255[37].9) OTU(MV_MV6R.CW.[CWD.MANDRV]) ] ,XIO(MV_N255[37].8) [OTU(MV_MV6R.CW.[CWD.MANUAL]) ,[XIC(MV_MV6R.CW.[CWD.OUTPUT]) OTL(MV_N255[37].9) ,XIO(MV_MV6R.CW.[CWD.OUTPUT]) OTU(MV_N255[37].9) ] ] ] ,[XIC(MV_N255[37].13) OTL(MV_MV6R.CW.[CWD.CHECKOFF]) ,XIO(MV_N255[37].13) OTU(MV_MV6R.CW.[CWD.CHECKOFF]) ] ] ,XIO(Delphi_Does_Eng_Func) [[XIC(MV_MV6R.CW.[CWD.MANUAL]) OTL(MV_N255[37].8) ,XIO(MV_MV6R.CW.[CWD.MANUAL]) OTU(MV_N255[37].8) ] ,[XIC(MV_MV6R.CW.[CWD.CHECKOFF]) OTL(MV_N255[37].13) ,XIO(MV_MV6R.CW.[CWD.CHECKOFF]) OTU(MV_N255[37].13) ] ,[XIC(MV_MV6R.CW.[CWD.OUTPUT]) OTL(MV_N255[37].9) ,XIO(MV_MV6R.CW.[CWD.OUTPUT]) OTU(MV_N255[37].9) ] ] ,XIC(MV_MV6R.CW.[CWD.RUNFB]) OTE(MV_N255[37].10) ,XIO(MV_MV6R.CW.[CWD.RUNFB]) OTE(MV_N255[37].11) ,XIC(MV_MV6R.CW.[CWD.FAULT]) OTE(MV_N255[37].15) ];
   47: [XIC(Delphi_Does_Eng_Func) [[XIC(MV_N255[38].8) [OTL(MV_MV7R.CW.[CWD.MANUAL]) ,XIC(MV_N255[38].9) OTL(MV_MV7R.CW.[CWD.MANDRV]) ,XIO(MV_N255[38].9) OTU(MV_MV7R.CW.[CWD.MANDRV]) ] ,XIO(MV_N255[38].8) [OTU(MV_MV7R.CW.[CWD.MANUAL]) ,[XIC(MV_MV7R.CW.[CWD.OUTPUT]) OTL(MV_N255[38].9) ,XIO(MV_MV7R.CW.[CWD.OUTPUT]) OTU(MV_N255[38].9) ] ] ] ,[XIC(MV_N255[38].13) OTL(MV_MV7R.CW.[CWD.CHECKOFF]) ,XIO(MV_N255[38].13) OTU(MV_MV7R.CW.[CWD.CHECKOFF]) ] ] ,XIO(Delphi_Does_Eng_Func) [[XIC(MV_MV7R.CW.[CWD.MANUAL]) OTL(MV_N255[38].8) ,XIO(MV_MV7R.CW.[CWD.MANUAL]) OTU(MV_N255[38].8) ] ,[XIC(MV_MV7R.CW.[CWD.CHECKOFF]) OTL(MV_N255[38].13) ,XIO(MV_MV7R.CW.[CWD.CHECKOFF]) OTU(MV_N255[38].13) ] ,[XIC(MV_MV7R.CW.[CWD.OUTPUT]) OTL(MV_N255[38].9) ,XIO(MV_MV7R.CW.[CWD.OUTPUT]) OTU(MV_N255[38].9) ] ] ,XIC(MV_MV7R.CW.[CWD.RUNFB]) OTE(MV_N255[38].10) ,XIO(MV_MV7R.CW.[CWD.RUNFB]) OTE(MV_N255[38].11) ,XIC(MV_MV7R.CW.[CWD.FAULT]) OTE(MV_N255[38].15) ];
